FUNCTION_BLOCK "FB100_Carrier"   // FB100, LAD
TITLE = Carrier Function Block
{ S7_Optimized_Access := 'TRUE' }
AUTHOR : INDICON
VERSION : 1.0
// Revision 1
   VAR_INPUT
      Position : DWord;
      CarrierNumber : Word;
      DriveStatus : "UDT_G120D_ZSW1_STATUS";
      DriveError : "UDT_G120D_ERRORS";
      DriveControlIn : "UDT_G120D_STW1_CONTROL";
      CommandSpeed : Word;
      ActualSpeedIn : Word;
      Reset : Bool;
      HMI : "UDT_CarrierHMI_In";
      PB_Box1_In : "UDT_PB_Box_In";
      PB_Box2_In : "UDT_PB_Box_In";
      SDC_In : "UDT_SDC_IN";
   END_VAR
   VAR_OUTPUT
      ReadyOn : Bool;
      Ready : Bool;
      Enabled : Bool;
      Stopped : Bool;
      MovingFwd : Bool;
      MovingREv : Bool;
      Fault : Bool;
      DriveControlOut : "UDT_G120D_STW1_CONTROL";
      CommandSpeedOut : Word;   // Control word output to Drive
      HMI_Out : "UDT_CarrierHMI_Out";
      Zone : Word;
      CarrierNUmConfirm : Word;
      CarrierPositionEcho : DWord;
      NextCarrierNum : Word;
      NextCarrierPos : Word;
      SDC_Out : "UDT_SDC_OUT";
      PB_Box1_Out : "UDT_PB_Box_Out";
      PB_Box2_Out : "UDT_PB_Box_Out";
   END_VAR
   VAR_TEMP
      DriveStatusTemp : Word;
      DriveControl_temp : "UDT_G120D_STW1_CONTROL";
      tempbit : Bool;
      tempbit1 : Bool;
      DriveStatusArray : "UDT_G120D_ZSW1_STATUS";
      Control_Out_Temp : "UDT_G120D_STW1_CONTROL";
      TempConversionFact : Real;
      ConversionFactor : Int;
   END_VAR
BEGIN

REGION Network 1: 1=EIN/ 0=AUS
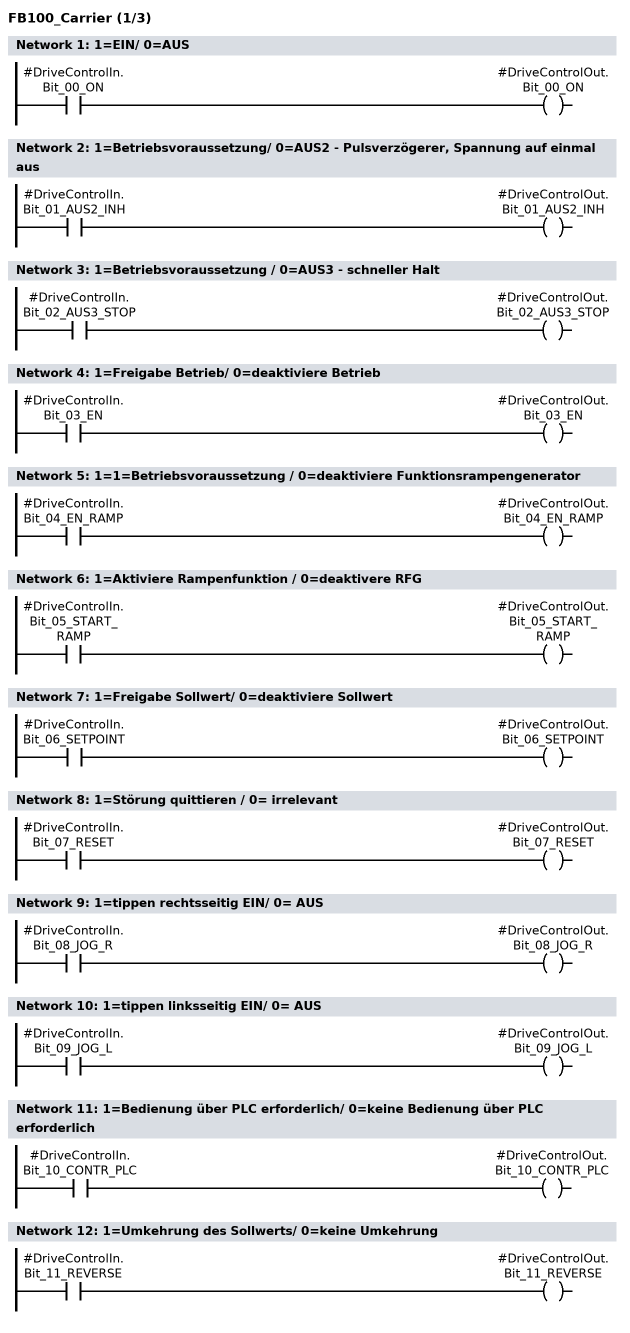
   RUNG wire#powerrail
      Contact( #DriveControlIn.Bit_00_ON )
      Coil( #DriveControlOut.Bit_00_ON )
   END_RUNG
   // the same network as SCL:
   #DriveControlOut.Bit_00_ON := #DriveControlIn.Bit_00_ON;
END_REGION

REGION Network 2: 1=Betriebsvoraussetzung/ 0=AUS2 - Pulsverzögerer, Spannung auf einmal aus
   RUNG wire#powerrail
      Contact( #DriveControlIn.Bit_01_AUS2_INH )
      Coil( #DriveControlOut.Bit_01_AUS2_INH )
   END_RUNG
   // the same network as SCL:
   #DriveControlOut.Bit_01_AUS2_INH := #DriveControlIn.Bit_01_AUS2_INH;
END_REGION

REGION Network 3: 1=Betriebsvoraussetzung / 0=AUS3 - schneller Halt
   RUNG wire#powerrail
      Contact( #DriveControlIn.Bit_02_AUS3_STOP )
      Coil( #DriveControlOut.Bit_02_AUS3_STOP )
   END_RUNG
   // the same network as SCL:
   #DriveControlOut.Bit_02_AUS3_STOP := #DriveControlIn.Bit_02_AUS3_STOP;
END_REGION

REGION Network 4: 1=Freigabe Betrieb/ 0=deaktiviere Betrieb
   RUNG wire#powerrail
      Contact( #DriveControlIn.Bit_03_EN )
      Coil( #DriveControlOut.Bit_03_EN )
   END_RUNG
   // the same network as SCL:
   #DriveControlOut.Bit_03_EN := #DriveControlIn.Bit_03_EN;
END_REGION

REGION Network 5: 1=1=Betriebsvoraussetzung / 0=deaktiviere Funktionsrampengenerator
   RUNG wire#powerrail
      Contact( #DriveControlIn.Bit_04_EN_RAMP )
      Coil( #DriveControlOut.Bit_04_EN_RAMP )
   END_RUNG
   // the same network as SCL:
   #DriveControlOut.Bit_04_EN_RAMP := #DriveControlIn.Bit_04_EN_RAMP;
END_REGION

REGION Network 6: 1=Aktiviere Rampenfunktion / 0=deaktivere RFG
   RUNG wire#powerrail
      Contact( #DriveControlIn.Bit_05_START_RAMP )
      Coil( #DriveControlOut.Bit_05_START_RAMP )
   END_RUNG
   // the same network as SCL:
   #DriveControlOut.Bit_05_START_RAMP := #DriveControlIn.Bit_05_START_RAMP;
END_REGION

REGION Network 7: 1=Freigabe Sollwert/ 0=deaktiviere Sollwert
   RUNG wire#powerrail
      Contact( #DriveControlIn.Bit_06_SETPOINT )
      Coil( #DriveControlOut.Bit_06_SETPOINT )
   END_RUNG
   // the same network as SCL:
   #DriveControlOut.Bit_06_SETPOINT := #DriveControlIn.Bit_06_SETPOINT;
END_REGION

REGION Network 8: 1=Störung quittieren / 0= irrelevant
   RUNG wire#powerrail
      Contact( #DriveControlIn.Bit_07_RESET )
      Coil( #DriveControlOut.Bit_07_RESET )
   END_RUNG
   // the same network as SCL:
   #DriveControlOut.Bit_07_RESET := #DriveControlIn.Bit_07_RESET;
END_REGION

REGION Network 9: 1=tippen rechtsseitig EIN/ 0= AUS
   RUNG wire#powerrail
      Contact( #DriveControlIn.Bit_08_JOG_R )
      Coil( #DriveControlOut.Bit_08_JOG_R )
   END_RUNG
   // the same network as SCL:
   #DriveControlOut.Bit_08_JOG_R := #DriveControlIn.Bit_08_JOG_R;
END_REGION

REGION Network 10: 1=tippen linksseitig EIN/ 0= AUS
   RUNG wire#powerrail
      Contact( #DriveControlIn.Bit_09_JOG_L )
      Coil( #DriveControlOut.Bit_09_JOG_L )
   END_RUNG
   // the same network as SCL:
   #DriveControlOut.Bit_09_JOG_L := #DriveControlIn.Bit_09_JOG_L;
END_REGION

REGION Network 11: 1=Bedienung über PLC erforderlich/ 0=keine Bedienung über PLC erforderlich
   RUNG wire#powerrail
      Contact( #DriveControlIn.Bit_10_CONTR_PLC )
      Coil( #DriveControlOut.Bit_10_CONTR_PLC )
   END_RUNG
   // the same network as SCL:
   #DriveControlOut.Bit_10_CONTR_PLC := #DriveControlIn.Bit_10_CONTR_PLC;
END_REGION

REGION Network 12: 1=Umkehrung des Sollwerts/ 0=keine Umkehrung
   RUNG wire#powerrail
      Contact( #DriveControlIn.Bit_11_REVERSE )
      Coil( #DriveControlOut.Bit_11_REVERSE )
   END_RUNG
   // the same network as SCL:
   #DriveControlOut.Bit_11_REVERSE := #DriveControlIn.Bit_11_REVERSE;
END_REGION

REGION Network 13: 1= Löse Bremse
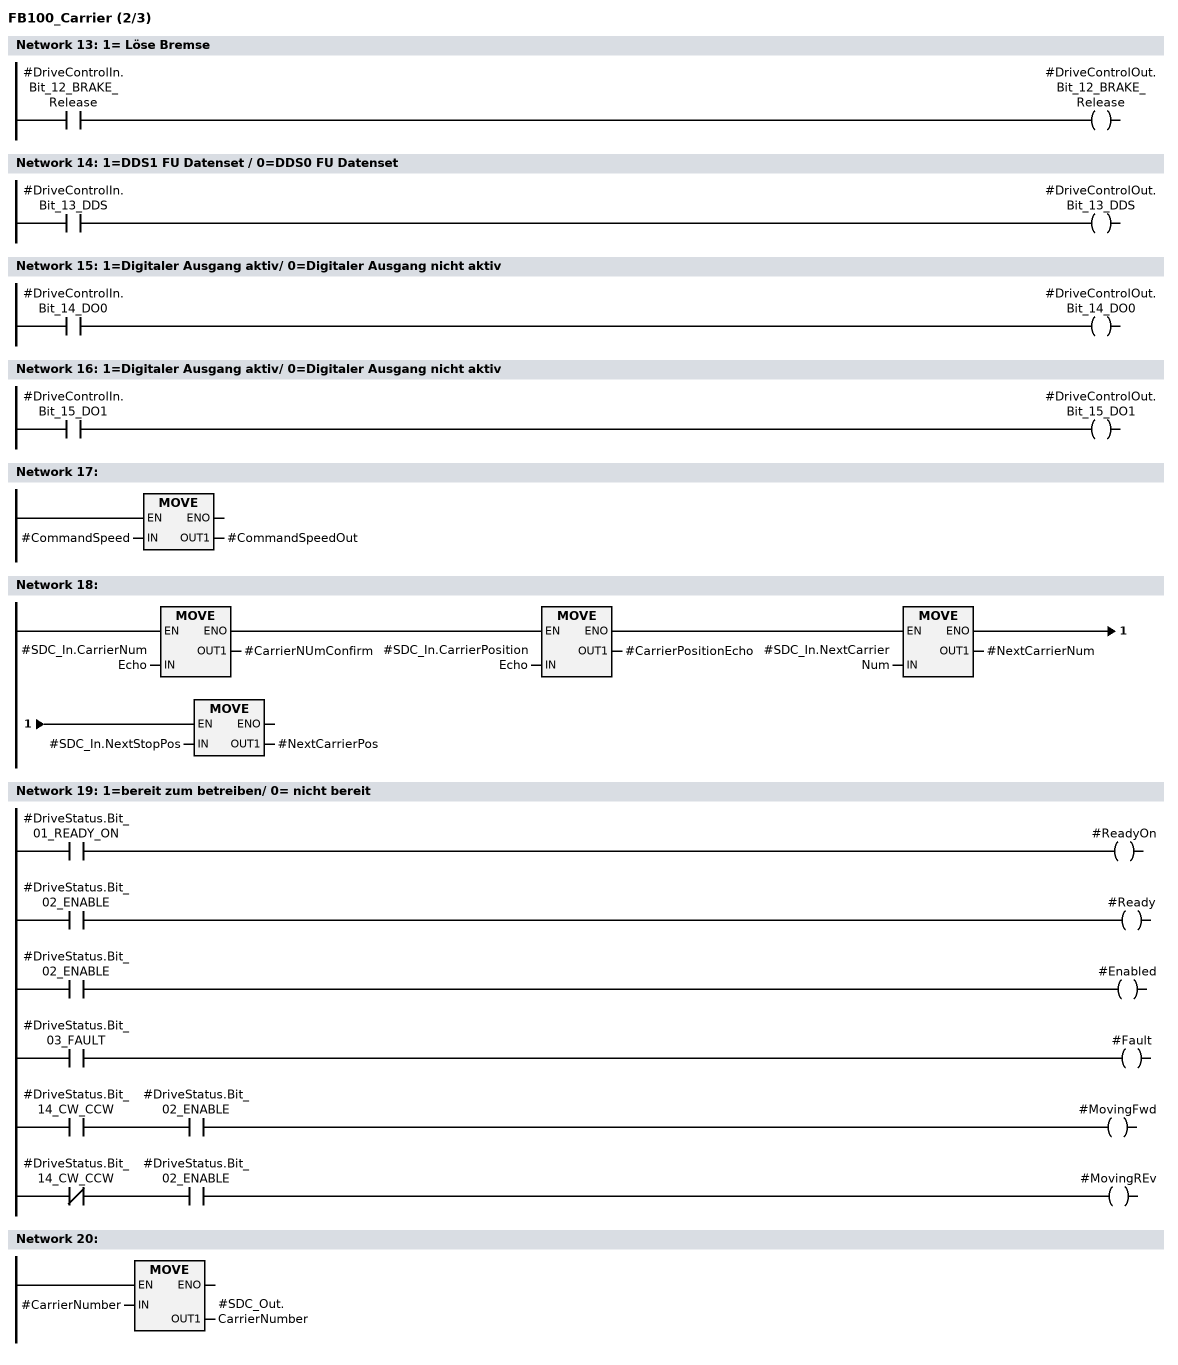
   RUNG wire#powerrail
      Contact( #DriveControlIn.Bit_12_BRAKE_Release )
      Coil( #DriveControlOut.Bit_12_BRAKE_Release )
   END_RUNG
   // the same network as SCL:
   #DriveControlOut.Bit_12_BRAKE_Release := #DriveControlIn.Bit_12_BRAKE_Release;
END_REGION

REGION Network 14: 1=DDS1 FU Datenset / 0=DDS0 FU Datenset
   RUNG wire#powerrail
      Contact( #DriveControlIn.Bit_13_DDS )
      Coil( #DriveControlOut.Bit_13_DDS )
   END_RUNG
   // the same network as SCL:
   #DriveControlOut.Bit_13_DDS := #DriveControlIn.Bit_13_DDS;
END_REGION

REGION Network 15: 1=Digitaler Ausgang aktiv/ 0=Digitaler Ausgang nicht aktiv
   RUNG wire#powerrail
      Contact( #DriveControlIn.Bit_14_DO0 )
      Coil( #DriveControlOut.Bit_14_DO0 )
   END_RUNG
   // the same network as SCL:
   #DriveControlOut.Bit_14_DO0 := #DriveControlIn.Bit_14_DO0;
END_REGION

REGION Network 16: 1=Digitaler Ausgang aktiv/ 0=Digitaler Ausgang nicht aktiv
   RUNG wire#powerrail
      Contact( #DriveControlIn.Bit_15_DO1 )
      Coil( #DriveControlOut.Bit_15_DO1 )
   END_RUNG
   // the same network as SCL:
   #DriveControlOut.Bit_15_DO1 := #DriveControlIn.Bit_15_DO1;
END_REGION

REGION Network 17
   RUNG wire#powerrail
      Move(in := #CommandSpeed, out1 => #CommandSpeedOut)
   END_RUNG
   // the same network as SCL:
   #CommandSpeedOut := #CommandSpeed;
END_REGION

REGION Network 18
   RUNG wire#powerrail
      Move(in := #SDC_In.CarrierNumEcho, out1 => #CarrierNUmConfirm)
      Move(in := #SDC_In.CarrierPositionEcho, out1 => #CarrierPositionEcho)
      Move(in := #SDC_In.NextCarrierNum, out1 => #NextCarrierNum)
      Move(in := #SDC_In.NextStopPos, out1 => #NextCarrierPos)
   END_RUNG
   // the same network as SCL:
   #CarrierNUmConfirm := #SDC_In.CarrierNumEcho;
   #CarrierPositionEcho := #SDC_In.CarrierPositionEcho;
   #NextCarrierNum := #SDC_In.NextCarrierNum;
   #NextCarrierPos := #SDC_In.NextStopPos;
END_REGION

REGION Network 19: 1=bereit zum betreiben/ 0= nicht bereit
   RUNG wire#powerrail
      Contact( #DriveStatus.Bit_01_READY_ON )
      Coil( #ReadyOn )
   END_RUNG
   RUNG wire#powerrail
      Contact( #DriveStatus.Bit_02_ENABLE )
      Coil( #Ready )
   END_RUNG
   RUNG wire#powerrail
      Contact( #DriveStatus.Bit_02_ENABLE )
      Coil( #Enabled )
   END_RUNG
   RUNG wire#powerrail
      Contact( #DriveStatus.Bit_03_FAULT )
      Coil( #Fault )
   END_RUNG
   RUNG wire#powerrail
      Contact( #DriveStatus.Bit_14_CW_CCW )
      Contact( #DriveStatus.Bit_02_ENABLE )
      Coil( #MovingFwd )
   END_RUNG
   RUNG wire#powerrail
      I_Contact( #DriveStatus.Bit_14_CW_CCW )
      Contact( #DriveStatus.Bit_02_ENABLE )
      Coil( #MovingREv )
   END_RUNG
   // the same network as SCL:
   #ReadyOn := #DriveStatus.Bit_01_READY_ON;
   #Ready := #DriveStatus.Bit_02_ENABLE;
   #Enabled := #DriveStatus.Bit_02_ENABLE;
   #Fault := #DriveStatus.Bit_03_FAULT;
   #MovingFwd := #DriveStatus.Bit_14_CW_CCW AND #DriveStatus.Bit_02_ENABLE;
   #MovingREv := NOT #DriveStatus.Bit_14_CW_CCW AND #DriveStatus.Bit_02_ENABLE;
END_REGION

REGION Network 20
   RUNG wire#powerrail
      Move(in := #CarrierNumber, out1 => #SDC_Out.CarrierNumber)
   END_RUNG
   // the same network as SCL:
   #SDC_Out.CarrierNumber := #CarrierNumber;
END_REGION

REGION Network 21
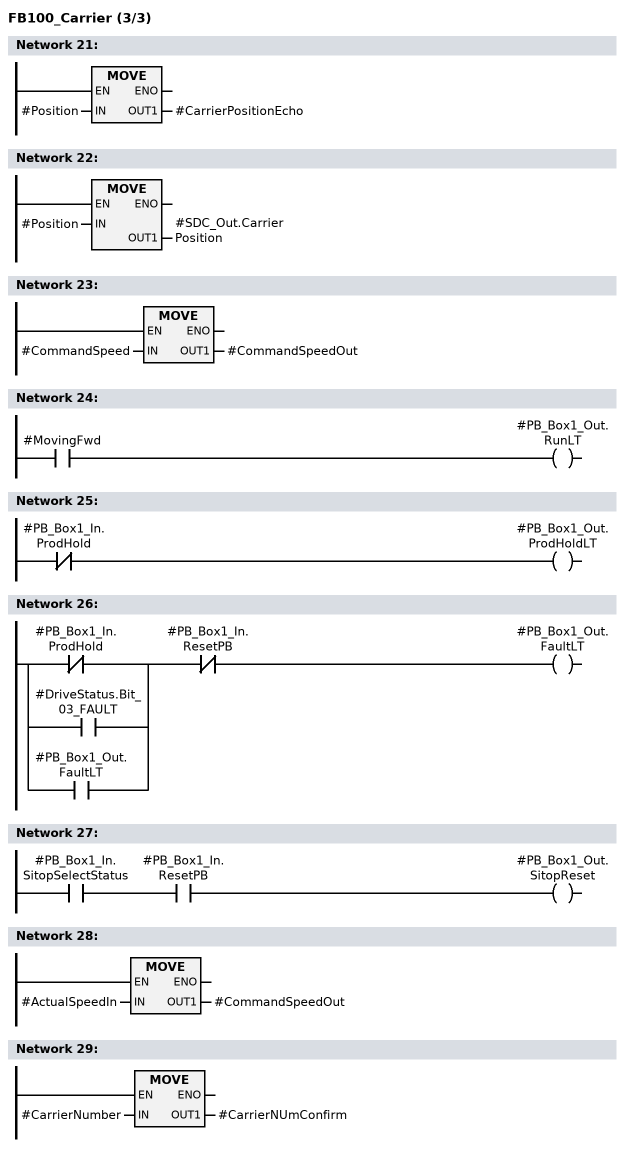
   RUNG wire#powerrail
      Move(in := #Position, out1 => #CarrierPositionEcho)
   END_RUNG
   // the same network as SCL:
   #CarrierPositionEcho := #Position;
END_REGION

REGION Network 22
   RUNG wire#powerrail
      Move(in := #Position, out1 => #SDC_Out.CarrierPosition)
   END_RUNG
   // the same network as SCL:
   #SDC_Out.CarrierPosition := #Position;
END_REGION

REGION Network 23
   RUNG wire#powerrail
      Move(in := #CommandSpeed, out1 => #CommandSpeedOut)
   END_RUNG
   // the same network as SCL:
   #CommandSpeedOut := #CommandSpeed;
END_REGION

REGION Network 24
   RUNG wire#powerrail
      Contact( #MovingFwd )
      Coil( #PB_Box1_Out.RunLT )
   END_RUNG
   // the same network as SCL:
   #PB_Box1_Out.RunLT := #MovingFwd;
END_REGION

REGION Network 25
   RUNG wire#powerrail
      I_Contact( #PB_Box1_In.ProdHold )
      Coil( #PB_Box1_Out.ProdHoldLT )
   END_RUNG
   // the same network as SCL:
   #PB_Box1_Out.ProdHoldLT := NOT #PB_Box1_In.ProdHold;
END_REGION

REGION Network 26
   RUNG wire#powerrail
      I_Contact( #PB_Box1_In.ProdHold )
      wire#w1
      I_Contact( #PB_Box1_In.ResetPB )
      Coil( #PB_Box1_Out.FaultLT )
   END_RUNG
   RUNG wire#powerrail
      Contact( #DriveStatus.Bit_03_FAULT )
   END_RUNG wire#w1
   RUNG wire#powerrail
      Contact( #PB_Box1_Out.FaultLT )
   END_RUNG wire#w1
   // the same network as SCL:
   #PB_Box1_Out.FaultLT := (NOT #PB_Box1_In.ProdHold OR #DriveStatus.Bit_03_FAULT OR #PB_Box1_Out.FaultLT) AND NOT #PB_Box1_In.ResetPB;
END_REGION

REGION Network 27
   RUNG wire#powerrail
      Contact( #PB_Box1_In.SitopSelectStatus )
      Contact( #PB_Box1_In.ResetPB )
      Coil( #PB_Box1_Out.SitopReset )
   END_RUNG
   // the same network as SCL:
   #PB_Box1_Out.SitopReset := #PB_Box1_In.SitopSelectStatus AND #PB_Box1_In.ResetPB;
END_REGION

REGION Network 28
   RUNG wire#powerrail
      Move(in := #ActualSpeedIn, out1 => #CommandSpeedOut)
   END_RUNG
   // the same network as SCL:
   #CommandSpeedOut := #ActualSpeedIn;
END_REGION

REGION Network 29
   RUNG wire#powerrail
      Move(in := #CarrierNumber, out1 => #CarrierNUmConfirm)
   END_RUNG
   // the same network as SCL:
   #CarrierNUmConfirm := #CarrierNumber;
END_REGION
END_FUNCTION_BLOCK

FUNCTION_BLOCK "FB101_ZONE"   // FB101, LAD
{ S7_Optimized_Access := 'TRUE' }
VERSION : 0.1
   VAR_INPUT
      ZONE : Int;
      DESCRIPTION : String;
      START_POSITION_IN : Int;
      END_POSITION_OUT : Int;
   END_VAR
   VAR_OUTPUT
      ZONE_ECHO : Int;
      START_POSITION : Int;
      STOP_POSITION : Int;
      DESCRIPTION_ECHO : String;
   END_VAR
BEGIN
END_FUNCTION_BLOCK

FUNCTION_BLOCK "FB102_Decode_Speed"   // FB102, LAD
{ S7_Optimized_Access := 'TRUE' }
VERSION : 0.1
   VAR_INPUT
      Speed : Word;
      Forward : Bool;
      Reverse : Bool;
   END_VAR
   VAR_OUTPUT
      Decimal1_Out : Word;
      Decimal2_Out : Word;
      Decimal3_Out : Word;
   END_VAR
   VAR RETAIN
      StringAll : String;
      String1 : String;
      String2 : String;
      String3 : String;
   END_VAR
   VAR_TEMP
      length : Word;
   END_VAR
BEGIN

REGION Network 1
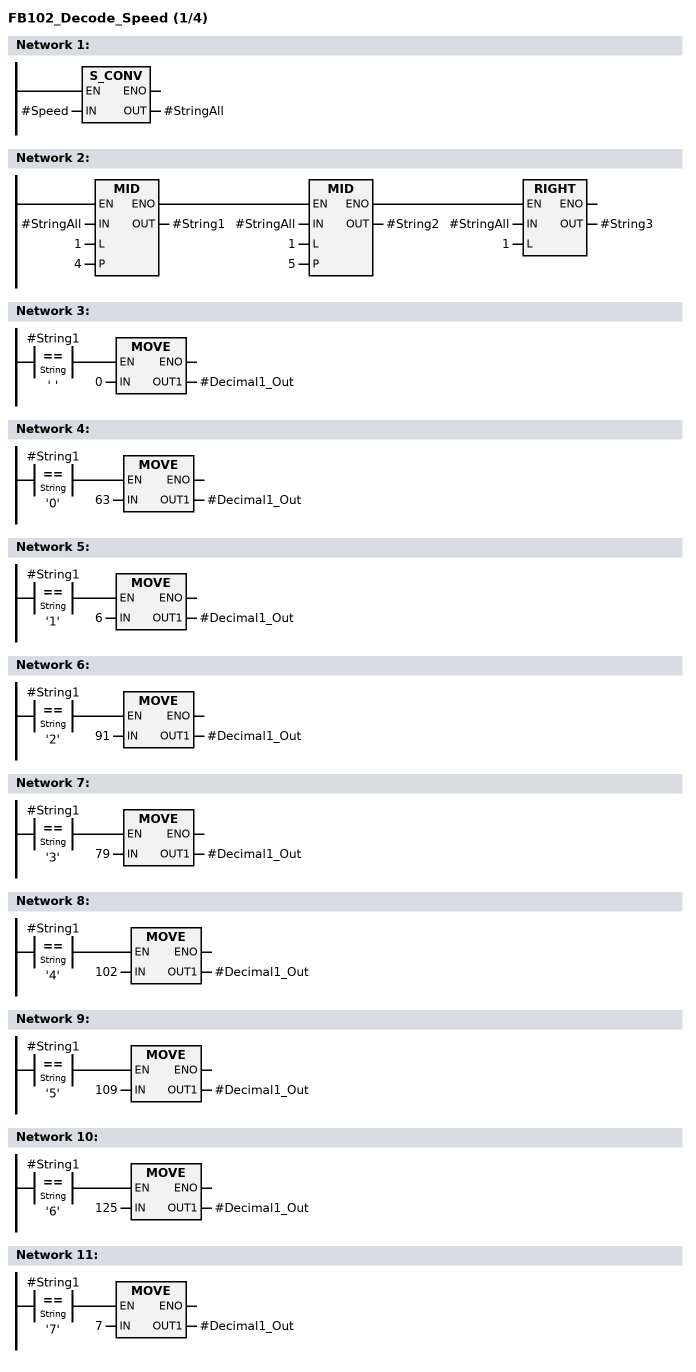
   #StringAll := S_CONV(IN := #Speed);
END_REGION

REGION Network 2
   #String1 := MID(IN := #StringAll, L := 1, P := 4);
   #String2 := MID(IN := #StringAll, L := 1, P := 5);
   #String3 := RIGHT(IN := #StringAll, L := 1);
END_REGION

REGION Network 3
   RUNG wire#powerrail
      { S7_Templates := "SrcType := String" } EQ_Contact(in1 := #String1, in2 := ' ')
      Move(in := 0, out1 => #Decimal1_Out)
   END_RUNG
   // the same network as SCL:
   IF #String1 = ' ' THEN #Decimal1_Out := 0; END_IF;
END_REGION

REGION Network 4
   RUNG wire#powerrail
      { S7_Templates := "SrcType := String" } EQ_Contact(in1 := #String1, in2 := '0')
      Move(in := 63, out1 => #Decimal1_Out)
   END_RUNG
   // the same network as SCL:
   IF #String1 = '0' THEN #Decimal1_Out := 63; END_IF;
END_REGION

REGION Network 5
   RUNG wire#powerrail
      { S7_Templates := "SrcType := String" } EQ_Contact(in1 := #String1, in2 := '1')
      Move(in := 6, out1 => #Decimal1_Out)
   END_RUNG
   // the same network as SCL:
   IF #String1 = '1' THEN #Decimal1_Out := 6; END_IF;
END_REGION

REGION Network 6
   RUNG wire#powerrail
      { S7_Templates := "SrcType := String" } EQ_Contact(in1 := #String1, in2 := '2')
      Move(in := 91, out1 => #Decimal1_Out)
   END_RUNG
   // the same network as SCL:
   IF #String1 = '2' THEN #Decimal1_Out := 91; END_IF;
END_REGION

REGION Network 7
   RUNG wire#powerrail
      { S7_Templates := "SrcType := String" } EQ_Contact(in1 := #String1, in2 := '3')
      Move(in := 79, out1 => #Decimal1_Out)
   END_RUNG
   // the same network as SCL:
   IF #String1 = '3' THEN #Decimal1_Out := 79; END_IF;
END_REGION

REGION Network 8
   RUNG wire#powerrail
      { S7_Templates := "SrcType := String" } EQ_Contact(in1 := #String1, in2 := '4')
      Move(in := 102, out1 => #Decimal1_Out)
   END_RUNG
   // the same network as SCL:
   IF #String1 = '4' THEN #Decimal1_Out := 102; END_IF;
END_REGION

REGION Network 9
   RUNG wire#powerrail
      { S7_Templates := "SrcType := String" } EQ_Contact(in1 := #String1, in2 := '5')
      Move(in := 109, out1 => #Decimal1_Out)
   END_RUNG
   // the same network as SCL:
   IF #String1 = '5' THEN #Decimal1_Out := 109; END_IF;
END_REGION

REGION Network 10
   RUNG wire#powerrail
      { S7_Templates := "SrcType := String" } EQ_Contact(in1 := #String1, in2 := '6')
      Move(in := 125, out1 => #Decimal1_Out)
   END_RUNG
   // the same network as SCL:
   IF #String1 = '6' THEN #Decimal1_Out := 125; END_IF;
END_REGION

REGION Network 11
   RUNG wire#powerrail
      { S7_Templates := "SrcType := String" } EQ_Contact(in1 := #String1, in2 := '7')
      Move(in := 7, out1 => #Decimal1_Out)
   END_RUNG
   // the same network as SCL:
   IF #String1 = '7' THEN #Decimal1_Out := 7; END_IF;
END_REGION

REGION Network 12
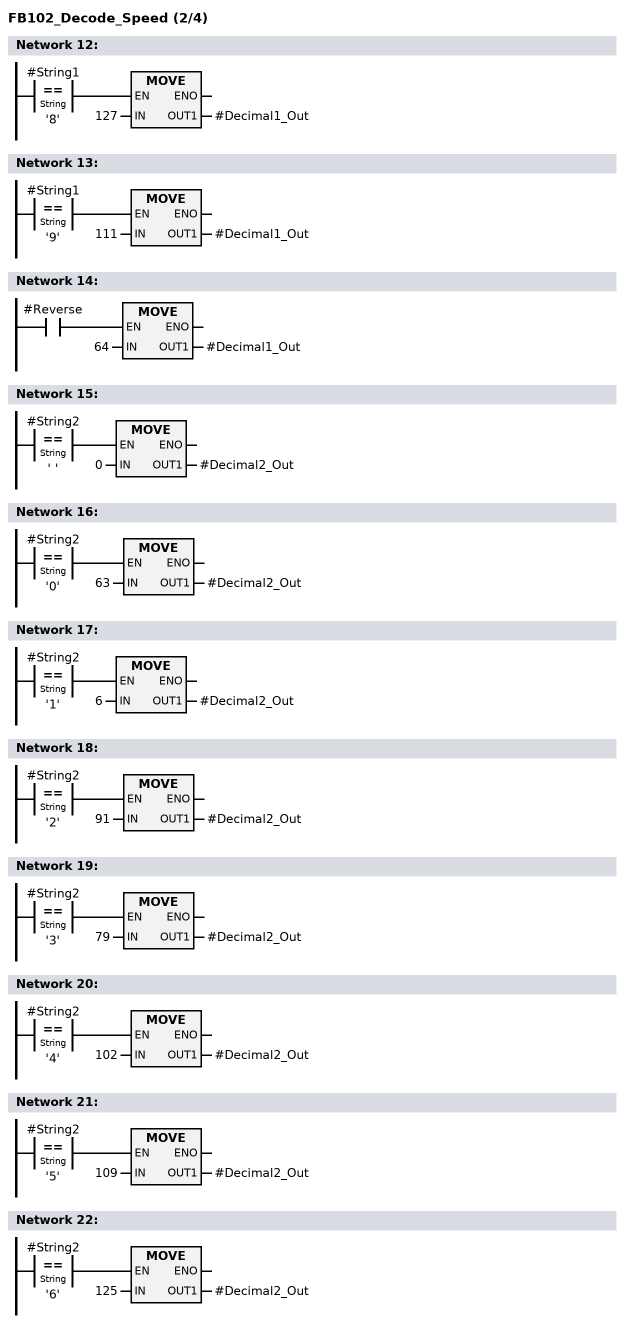
   RUNG wire#powerrail
      { S7_Templates := "SrcType := String" } EQ_Contact(in1 := #String1, in2 := '8')
      Move(in := 127, out1 => #Decimal1_Out)
   END_RUNG
   // the same network as SCL:
   IF #String1 = '8' THEN #Decimal1_Out := 127; END_IF;
END_REGION

REGION Network 13
   RUNG wire#powerrail
      { S7_Templates := "SrcType := String" } EQ_Contact(in1 := #String1, in2 := '9')
      Move(in := 111, out1 => #Decimal1_Out)
   END_RUNG
   // the same network as SCL:
   IF #String1 = '9' THEN #Decimal1_Out := 111; END_IF;
END_REGION

REGION Network 14
   RUNG wire#powerrail
      Contact( #Reverse )
      Move(in := 64, out1 => #Decimal1_Out)
   END_RUNG
   // the same network as SCL:
   IF #Reverse THEN #Decimal1_Out := 64; END_IF;
END_REGION

REGION Network 15
   RUNG wire#powerrail
      { S7_Templates := "SrcType := String" } EQ_Contact(in1 := #String2, in2 := ' ')
      Move(in := 0, out1 => #Decimal2_Out)
   END_RUNG
   // the same network as SCL:
   IF #String2 = ' ' THEN #Decimal2_Out := 0; END_IF;
END_REGION

REGION Network 16
   RUNG wire#powerrail
      { S7_Templates := "SrcType := String" } EQ_Contact(in1 := #String2, in2 := '0')
      Move(in := 63, out1 => #Decimal2_Out)
   END_RUNG
   // the same network as SCL:
   IF #String2 = '0' THEN #Decimal2_Out := 63; END_IF;
END_REGION

REGION Network 17
   RUNG wire#powerrail
      { S7_Templates := "SrcType := String" } EQ_Contact(in1 := #String2, in2 := '1')
      Move(in := 6, out1 => #Decimal2_Out)
   END_RUNG
   // the same network as SCL:
   IF #String2 = '1' THEN #Decimal2_Out := 6; END_IF;
END_REGION

REGION Network 18
   RUNG wire#powerrail
      { S7_Templates := "SrcType := String" } EQ_Contact(in1 := #String2, in2 := '2')
      Move(in := 91, out1 => #Decimal2_Out)
   END_RUNG
   // the same network as SCL:
   IF #String2 = '2' THEN #Decimal2_Out := 91; END_IF;
END_REGION

REGION Network 19
   RUNG wire#powerrail
      { S7_Templates := "SrcType := String" } EQ_Contact(in1 := #String2, in2 := '3')
      Move(in := 79, out1 => #Decimal2_Out)
   END_RUNG
   // the same network as SCL:
   IF #String2 = '3' THEN #Decimal2_Out := 79; END_IF;
END_REGION

REGION Network 20
   RUNG wire#powerrail
      { S7_Templates := "SrcType := String" } EQ_Contact(in1 := #String2, in2 := '4')
      Move(in := 102, out1 => #Decimal2_Out)
   END_RUNG
   // the same network as SCL:
   IF #String2 = '4' THEN #Decimal2_Out := 102; END_IF;
END_REGION

REGION Network 21
   RUNG wire#powerrail
      { S7_Templates := "SrcType := String" } EQ_Contact(in1 := #String2, in2 := '5')
      Move(in := 109, out1 => #Decimal2_Out)
   END_RUNG
   // the same network as SCL:
   IF #String2 = '5' THEN #Decimal2_Out := 109; END_IF;
END_REGION

REGION Network 22
   RUNG wire#powerrail
      { S7_Templates := "SrcType := String" } EQ_Contact(in1 := #String2, in2 := '6')
      Move(in := 125, out1 => #Decimal2_Out)
   END_RUNG
   // the same network as SCL:
   IF #String2 = '6' THEN #Decimal2_Out := 125; END_IF;
END_REGION

REGION Network 23
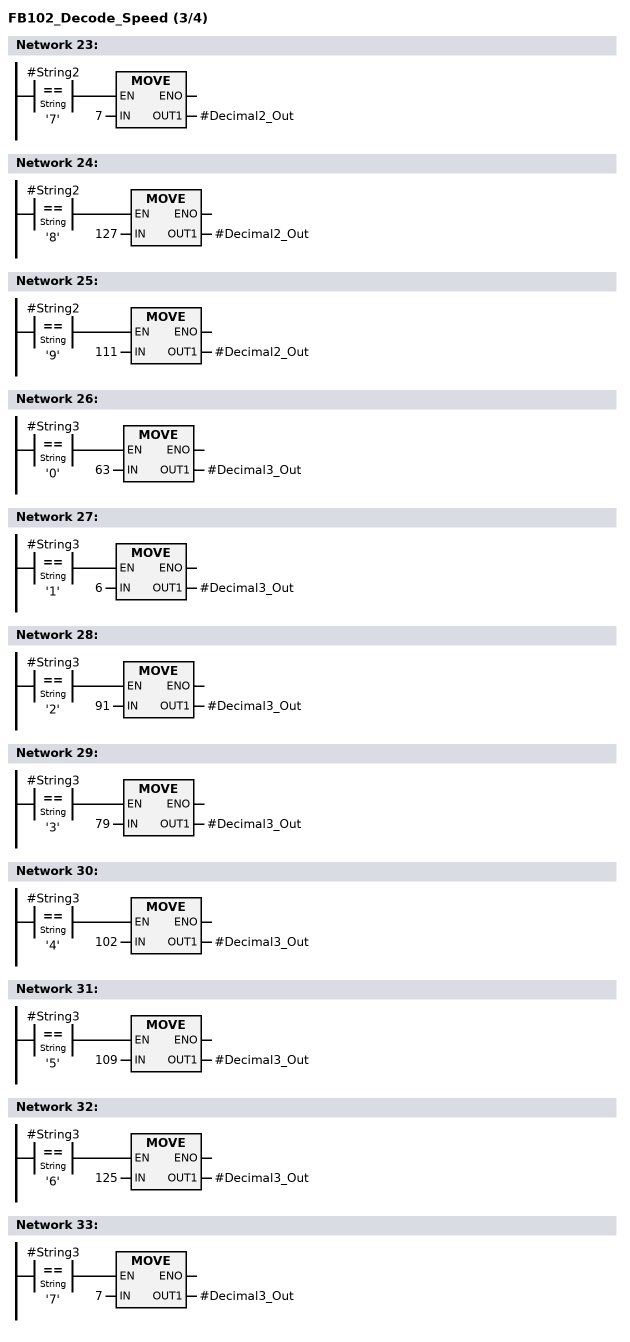
   RUNG wire#powerrail
      { S7_Templates := "SrcType := String" } EQ_Contact(in1 := #String2, in2 := '7')
      Move(in := 7, out1 => #Decimal2_Out)
   END_RUNG
   // the same network as SCL:
   IF #String2 = '7' THEN #Decimal2_Out := 7; END_IF;
END_REGION

REGION Network 24
   RUNG wire#powerrail
      { S7_Templates := "SrcType := String" } EQ_Contact(in1 := #String2, in2 := '8')
      Move(in := 127, out1 => #Decimal2_Out)
   END_RUNG
   // the same network as SCL:
   IF #String2 = '8' THEN #Decimal2_Out := 127; END_IF;
END_REGION

REGION Network 25
   RUNG wire#powerrail
      { S7_Templates := "SrcType := String" } EQ_Contact(in1 := #String2, in2 := '9')
      Move(in := 111, out1 => #Decimal2_Out)
   END_RUNG
   // the same network as SCL:
   IF #String2 = '9' THEN #Decimal2_Out := 111; END_IF;
END_REGION

REGION Network 26
   RUNG wire#powerrail
      { S7_Templates := "SrcType := String" } EQ_Contact(in1 := #String3, in2 := '0')
      Move(in := 63, out1 => #Decimal3_Out)
   END_RUNG
   // the same network as SCL:
   IF #String3 = '0' THEN #Decimal3_Out := 63; END_IF;
END_REGION

REGION Network 27
   RUNG wire#powerrail
      { S7_Templates := "SrcType := String" } EQ_Contact(in1 := #String3, in2 := '1')
      Move(in := 6, out1 => #Decimal3_Out)
   END_RUNG
   // the same network as SCL:
   IF #String3 = '1' THEN #Decimal3_Out := 6; END_IF;
END_REGION

REGION Network 28
   RUNG wire#powerrail
      { S7_Templates := "SrcType := String" } EQ_Contact(in1 := #String3, in2 := '2')
      Move(in := 91, out1 => #Decimal3_Out)
   END_RUNG
   // the same network as SCL:
   IF #String3 = '2' THEN #Decimal3_Out := 91; END_IF;
END_REGION

REGION Network 29
   RUNG wire#powerrail
      { S7_Templates := "SrcType := String" } EQ_Contact(in1 := #String3, in2 := '3')
      Move(in := 79, out1 => #Decimal3_Out)
   END_RUNG
   // the same network as SCL:
   IF #String3 = '3' THEN #Decimal3_Out := 79; END_IF;
END_REGION

REGION Network 30
   RUNG wire#powerrail
      { S7_Templates := "SrcType := String" } EQ_Contact(in1 := #String3, in2 := '4')
      Move(in := 102, out1 => #Decimal3_Out)
   END_RUNG
   // the same network as SCL:
   IF #String3 = '4' THEN #Decimal3_Out := 102; END_IF;
END_REGION

REGION Network 31
   RUNG wire#powerrail
      { S7_Templates := "SrcType := String" } EQ_Contact(in1 := #String3, in2 := '5')
      Move(in := 109, out1 => #Decimal3_Out)
   END_RUNG
   // the same network as SCL:
   IF #String3 = '5' THEN #Decimal3_Out := 109; END_IF;
END_REGION

REGION Network 32
   RUNG wire#powerrail
      { S7_Templates := "SrcType := String" } EQ_Contact(in1 := #String3, in2 := '6')
      Move(in := 125, out1 => #Decimal3_Out)
   END_RUNG
   // the same network as SCL:
   IF #String3 = '6' THEN #Decimal3_Out := 125; END_IF;
END_REGION

REGION Network 33
   RUNG wire#powerrail
      { S7_Templates := "SrcType := String" } EQ_Contact(in1 := #String3, in2 := '7')
      Move(in := 7, out1 => #Decimal3_Out)
   END_RUNG
   // the same network as SCL:
   IF #String3 = '7' THEN #Decimal3_Out := 7; END_IF;
END_REGION

REGION Network 34
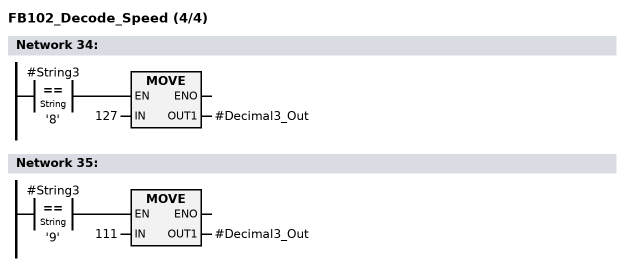
   RUNG wire#powerrail
      { S7_Templates := "SrcType := String" } EQ_Contact(in1 := #String3, in2 := '8')
      Move(in := 127, out1 => #Decimal3_Out)
   END_RUNG
   // the same network as SCL:
   IF #String3 = '8' THEN #Decimal3_Out := 127; END_IF;
END_REGION

REGION Network 35
   RUNG wire#powerrail
      { S7_Templates := "SrcType := String" } EQ_Contact(in1 := #String3, in2 := '9')
      Move(in := 111, out1 => #Decimal3_Out)
   END_RUNG
   // the same network as SCL:
   IF #String3 = '9' THEN #Decimal3_Out := 111; END_IF;
END_REGION
END_FUNCTION_BLOCK

FUNCTION_BLOCK "FB103_Decode_Carrier_Number"   // FB103, LAD
{ S7_Optimized_Access := 'TRUE' }
VERSION : 0.1
   VAR_INPUT
      Carrier_Number : Word;
   END_VAR
   VAR_OUTPUT
      Decimal1_Out : Word;
      Decimal2_Out : Word;
      Decimal3_Out : Word;
   END_VAR
   VAR RETAIN
      StringAll : String;
      String1 : String;
      String2 : String;
      String3 : String;
   END_VAR
   VAR_TEMP
      length : Word;
   END_VAR
BEGIN

REGION Network 1
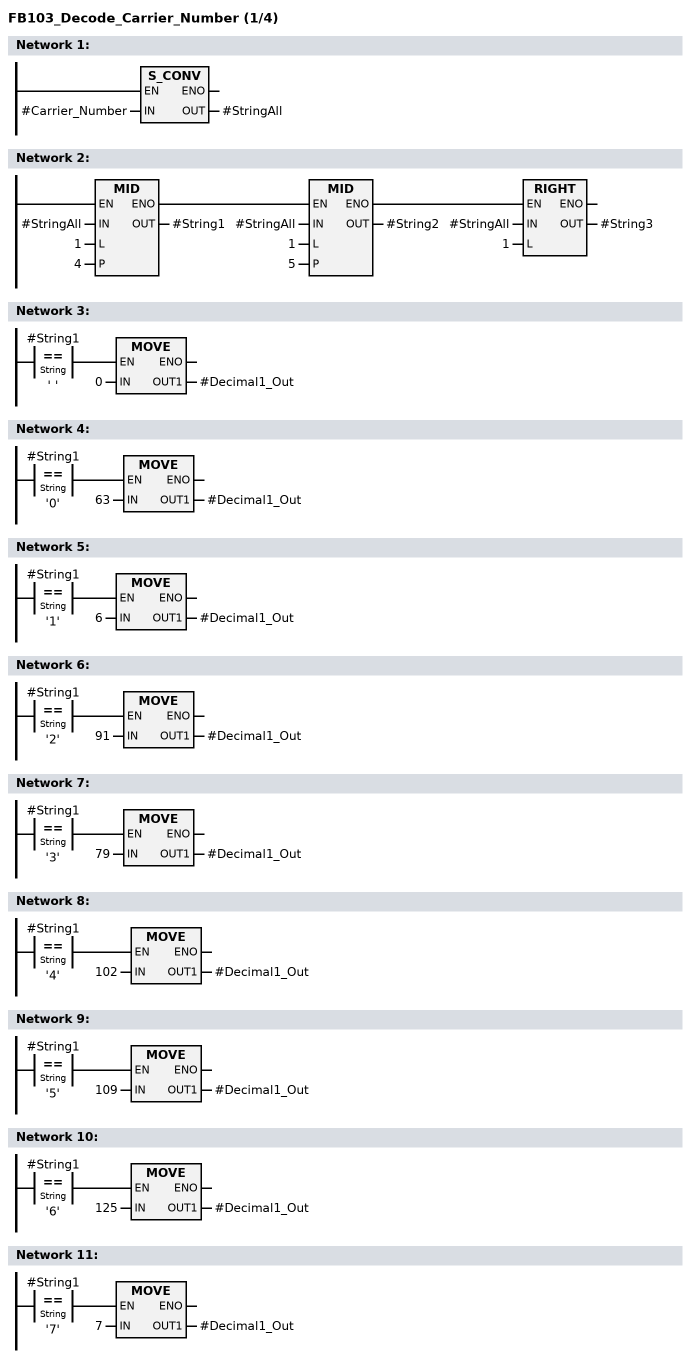
   #StringAll := S_CONV(IN := #Carrier_Number);
END_REGION

REGION Network 2
   #String1 := MID(IN := #StringAll, L := 1, P := 4);
   #String2 := MID(IN := #StringAll, L := 1, P := 5);
   #String3 := RIGHT(IN := #StringAll, L := 1);
END_REGION

REGION Network 3
   RUNG wire#powerrail
      { S7_Templates := "SrcType := String" } EQ_Contact(in1 := #String1, in2 := ' ')
      Move(in := 0, out1 => #Decimal1_Out)
   END_RUNG
   // the same network as SCL:
   IF #String1 = ' ' THEN #Decimal1_Out := 0; END_IF;
END_REGION

REGION Network 4
   RUNG wire#powerrail
      { S7_Templates := "SrcType := String" } EQ_Contact(in1 := #String1, in2 := '0')
      Move(in := 63, out1 => #Decimal1_Out)
   END_RUNG
   // the same network as SCL:
   IF #String1 = '0' THEN #Decimal1_Out := 63; END_IF;
END_REGION

REGION Network 5
   RUNG wire#powerrail
      { S7_Templates := "SrcType := String" } EQ_Contact(in1 := #String1, in2 := '1')
      Move(in := 6, out1 => #Decimal1_Out)
   END_RUNG
   // the same network as SCL:
   IF #String1 = '1' THEN #Decimal1_Out := 6; END_IF;
END_REGION

REGION Network 6
   RUNG wire#powerrail
      { S7_Templates := "SrcType := String" } EQ_Contact(in1 := #String1, in2 := '2')
      Move(in := 91, out1 => #Decimal1_Out)
   END_RUNG
   // the same network as SCL:
   IF #String1 = '2' THEN #Decimal1_Out := 91; END_IF;
END_REGION

REGION Network 7
   RUNG wire#powerrail
      { S7_Templates := "SrcType := String" } EQ_Contact(in1 := #String1, in2 := '3')
      Move(in := 79, out1 => #Decimal1_Out)
   END_RUNG
   // the same network as SCL:
   IF #String1 = '3' THEN #Decimal1_Out := 79; END_IF;
END_REGION

REGION Network 8
   RUNG wire#powerrail
      { S7_Templates := "SrcType := String" } EQ_Contact(in1 := #String1, in2 := '4')
      Move(in := 102, out1 => #Decimal1_Out)
   END_RUNG
   // the same network as SCL:
   IF #String1 = '4' THEN #Decimal1_Out := 102; END_IF;
END_REGION

REGION Network 9
   RUNG wire#powerrail
      { S7_Templates := "SrcType := String" } EQ_Contact(in1 := #String1, in2 := '5')
      Move(in := 109, out1 => #Decimal1_Out)
   END_RUNG
   // the same network as SCL:
   IF #String1 = '5' THEN #Decimal1_Out := 109; END_IF;
END_REGION

REGION Network 10
   RUNG wire#powerrail
      { S7_Templates := "SrcType := String" } EQ_Contact(in1 := #String1, in2 := '6')
      Move(in := 125, out1 => #Decimal1_Out)
   END_RUNG
   // the same network as SCL:
   IF #String1 = '6' THEN #Decimal1_Out := 125; END_IF;
END_REGION

REGION Network 11
   RUNG wire#powerrail
      { S7_Templates := "SrcType := String" } EQ_Contact(in1 := #String1, in2 := '7')
      Move(in := 7, out1 => #Decimal1_Out)
   END_RUNG
   // the same network as SCL:
   IF #String1 = '7' THEN #Decimal1_Out := 7; END_IF;
END_REGION

REGION Network 12
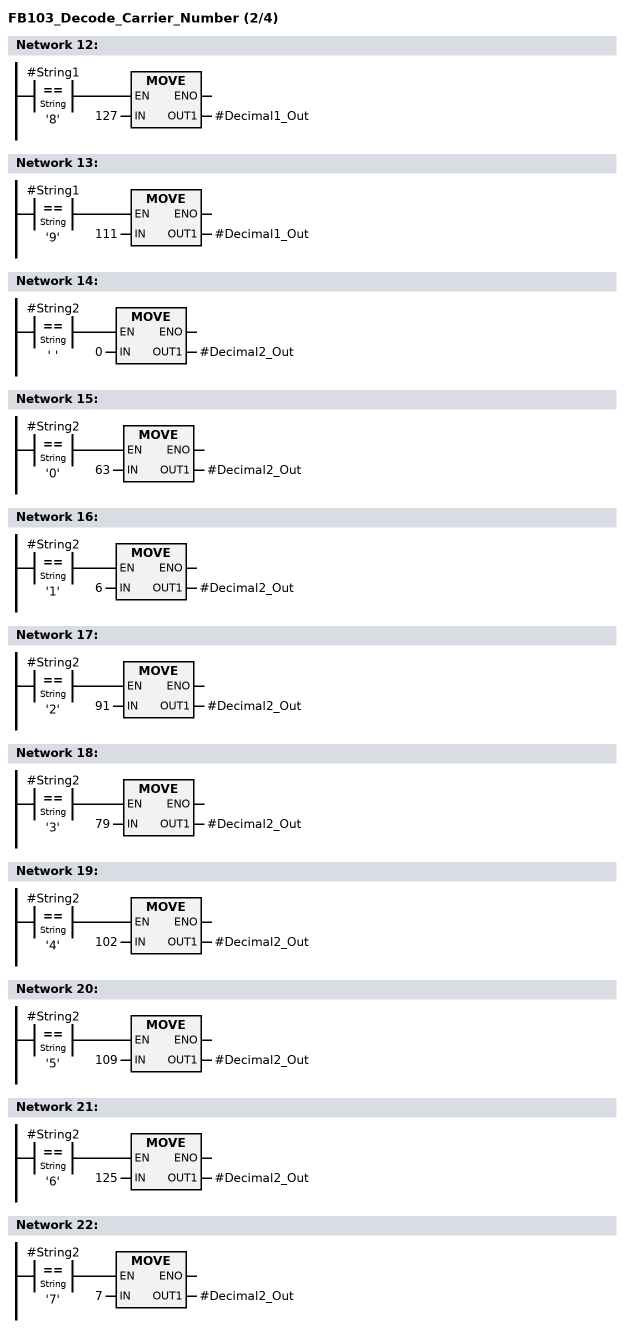
   RUNG wire#powerrail
      { S7_Templates := "SrcType := String" } EQ_Contact(in1 := #String1, in2 := '8')
      Move(in := 127, out1 => #Decimal1_Out)
   END_RUNG
   // the same network as SCL:
   IF #String1 = '8' THEN #Decimal1_Out := 127; END_IF;
END_REGION

REGION Network 13
   RUNG wire#powerrail
      { S7_Templates := "SrcType := String" } EQ_Contact(in1 := #String1, in2 := '9')
      Move(in := 111, out1 => #Decimal1_Out)
   END_RUNG
   // the same network as SCL:
   IF #String1 = '9' THEN #Decimal1_Out := 111; END_IF;
END_REGION

REGION Network 14
   RUNG wire#powerrail
      { S7_Templates := "SrcType := String" } EQ_Contact(in1 := #String2, in2 := ' ')
      Move(in := 0, out1 => #Decimal2_Out)
   END_RUNG
   // the same network as SCL:
   IF #String2 = ' ' THEN #Decimal2_Out := 0; END_IF;
END_REGION

REGION Network 15
   RUNG wire#powerrail
      { S7_Templates := "SrcType := String" } EQ_Contact(in1 := #String2, in2 := '0')
      Move(in := 63, out1 => #Decimal2_Out)
   END_RUNG
   // the same network as SCL:
   IF #String2 = '0' THEN #Decimal2_Out := 63; END_IF;
END_REGION

REGION Network 16
   RUNG wire#powerrail
      { S7_Templates := "SrcType := String" } EQ_Contact(in1 := #String2, in2 := '1')
      Move(in := 6, out1 => #Decimal2_Out)
   END_RUNG
   // the same network as SCL:
   IF #String2 = '1' THEN #Decimal2_Out := 6; END_IF;
END_REGION

REGION Network 17
   RUNG wire#powerrail
      { S7_Templates := "SrcType := String" } EQ_Contact(in1 := #String2, in2 := '2')
      Move(in := 91, out1 => #Decimal2_Out)
   END_RUNG
   // the same network as SCL:
   IF #String2 = '2' THEN #Decimal2_Out := 91; END_IF;
END_REGION

REGION Network 18
   RUNG wire#powerrail
      { S7_Templates := "SrcType := String" } EQ_Contact(in1 := #String2, in2 := '3')
      Move(in := 79, out1 => #Decimal2_Out)
   END_RUNG
   // the same network as SCL:
   IF #String2 = '3' THEN #Decimal2_Out := 79; END_IF;
END_REGION

REGION Network 19
   RUNG wire#powerrail
      { S7_Templates := "SrcType := String" } EQ_Contact(in1 := #String2, in2 := '4')
      Move(in := 102, out1 => #Decimal2_Out)
   END_RUNG
   // the same network as SCL:
   IF #String2 = '4' THEN #Decimal2_Out := 102; END_IF;
END_REGION

REGION Network 20
   RUNG wire#powerrail
      { S7_Templates := "SrcType := String" } EQ_Contact(in1 := #String2, in2 := '5')
      Move(in := 109, out1 => #Decimal2_Out)
   END_RUNG
   // the same network as SCL:
   IF #String2 = '5' THEN #Decimal2_Out := 109; END_IF;
END_REGION
